REGION Network 46: Aviso 55 - El Secador Sullair 1 alcanzó la máxima cantidad de horas sin mantenimiento 2
   RUNG wire#powerrail
      Contact( "LimiteMantMS054_2" )
      Coil( "DB_ALA_PRE".x165 )
   END_RUNG
   // the same network as SCL:
   "DB_ALA_PRE".x165 := "LimiteMantMS054_2";
END_REGION

REGION Network 47: Aviso 56 - El Secador Sullair 2 alcanzó la máxima cantidad de horas sin mantenimiento 1
   RUNG wire#powerrail
      Contact( "LimiteMantMS055_1" )
      Coil( "DB_ALA_PRE".x166 )
   END_RUNG
   // the same network as SCL:
   "DB_ALA_PRE".x166 := "LimiteMantMS055_1";
END_REGION

REGION Network 48: Aviso 57 - El Secador Sullair 2 alcanzó la máxima cantidad de horas sin mantenimiento 2
   RUNG wire#powerrail
      Contact( "LimiteMantMS055_2" )
      Coil( "DB_ALA_PRE".x167 )
   END_RUNG
   // the same network as SCL:
   "DB_ALA_PRE".x167 := "LimiteMantMS055_2";
END_REGION

REGION Network 49: Aviso 58 - El Compresor Sullair 2 alcanzó la máxima cantidad de horas sin mantenimiento 1
   RUNG wire#powerrail
      Contact( "LimiteMantMC060_1" )
      Coil( "DB_ALA_PRE".x168 )
   END_RUNG
   // the same network as SCL:
   "DB_ALA_PRE".x168 := "LimiteMantMC060_1";
END_REGION

REGION Network 50: Aviso 59 - El Compresor Sullair 2 alcanzó la máxima cantidad de horas sin mantenimiento 2
   RUNG wire#powerrail
      Contact( "LimiteMantMC060_2" )
      Coil( "DB_ALA_PRE".x169 )
   END_RUNG
   // the same network as SCL:
   "DB_ALA_PRE".x169 := "LimiteMantMC060_2";
END_REGION

REGION Network 51: Aviso 60 - El Compresor Sullair 2 alcanzó la máxima cantidad de horas sin mantenimiento 3
   RUNG wire#powerrail
      Contact( "LimiteMantMC060_3" )
      Coil( "DB_ALA_PRE".x170 )
   END_RUNG
   // the same network as SCL:
   "DB_ALA_PRE".x170 := "LimiteMantMC060_3";
END_REGION

REGION Network 52: Aviso 61 - El Compresor Sullair 2 alcanzó la máxima cantidad de horas sin mantenimiento 4
   RUNG wire#powerrail
      Contact( "LimiteMantMC060_4" )
      Coil( "DB_ALA_PRE".x171 )
   END_RUNG
   // the same network as SCL:
   "DB_ALA_PRE".x171 := "LimiteMantMC060_4";
END_REGION

REGION Network 53: Aviso 62 - El Compresor Sullair 2 alcanzó la máxima cantidad de horas sin mantenimiento 5
   RUNG wire#powerrail
      Contact( "LimiteMantMC060_5" )
      Coil( "DB_ALA_PRE".x172 )
   END_RUNG
   // the same network as SCL:
   "DB_ALA_PRE".x172 := "LimiteMantMC060_5";
END_REGION

REGION Network 54: Aviso 63 - El Compresor Sullair 1 alcanzó la máxima cantidad de horas sin mantenimiento 1
   RUNG wire#powerrail
      Contact( "LimiteMantMC061_1" )
      Coil( "DB_ALA_PRE".x173 )
   END_RUNG
   // the same network as SCL:
   "DB_ALA_PRE".x173 := "LimiteMantMC061_1";
END_REGION

REGION Network 55: Aviso 64 - El Compresor Sullair 1 alcanzó la máxima cantidad de horas sin mantenimiento 2
   RUNG wire#powerrail
      Contact( "LimiteMantMC061_2" )
      Coil( "DB_ALA_PRE".x174 )
   END_RUNG
   // the same network as SCL:
   "DB_ALA_PRE".x174 := "LimiteMantMC061_2";
END_REGION

REGION Network 56: Aviso 65 - El Compresor Sullair 1 alcanzó la máxima cantidad de horas sin mantenimiento 3
   RUNG wire#powerrail
      Contact( "LimiteMantMC061_3" )
      Coil( "DB_ALA_PRE".x175 )
   END_RUNG
   // the same network as SCL:
   "DB_ALA_PRE".x175 := "LimiteMantMC061_3";
END_REGION

REGION Network 57: Aviso 84 - El Compresor Sullair 1 alcanzó la máxima cantidad de horas sin mantenimiento 4
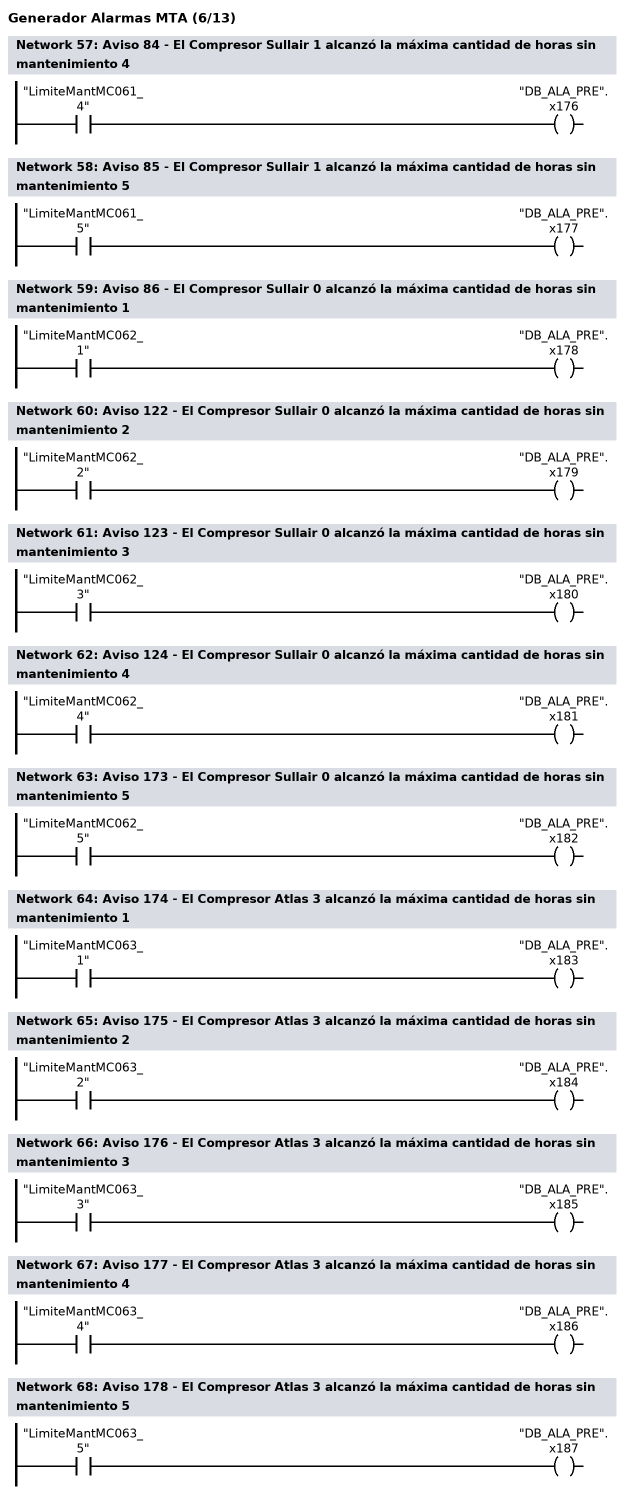
   RUNG wire#powerrail
      Contact( "LimiteMantMC061_4" )
      Coil( "DB_ALA_PRE".x176 )
   END_RUNG
   // the same network as SCL:
   "DB_ALA_PRE".x176 := "LimiteMantMC061_4";
END_REGION

REGION Network 58: Aviso 85 - El Compresor Sullair 1 alcanzó la máxima cantidad de horas sin mantenimiento 5
   RUNG wire#powerrail
      Contact( "LimiteMantMC061_5" )
      Coil( "DB_ALA_PRE".x177 )
   END_RUNG
   // the same network as SCL:
   "DB_ALA_PRE".x177 := "LimiteMantMC061_5";
END_REGION

REGION Network 59: Aviso 86 - El Compresor Sullair 0 alcanzó la máxima cantidad de horas sin mantenimiento 1
   RUNG wire#powerrail
      Contact( "LimiteMantMC062_1" )
      Coil( "DB_ALA_PRE".x178 )
   END_RUNG
   // the same network as SCL:
   "DB_ALA_PRE".x178 := "LimiteMantMC062_1";
END_REGION

REGION Network 60: Aviso 122 - El Compresor Sullair 0 alcanzó la máxima cantidad de horas sin mantenimiento 2
   RUNG wire#powerrail
      Contact( "LimiteMantMC062_2" )
      Coil( "DB_ALA_PRE".x179 )
   END_RUNG
   // the same network as SCL:
   "DB_ALA_PRE".x179 := "LimiteMantMC062_2";
END_REGION

REGION Network 61: Aviso 123 - El Compresor Sullair 0 alcanzó la máxima cantidad de horas sin mantenimiento 3
   RUNG wire#powerrail
      Contact( "LimiteMantMC062_3" )
      Coil( "DB_ALA_PRE".x180 )
   END_RUNG
   // the same network as SCL:
   "DB_ALA_PRE".x180 := "LimiteMantMC062_3";
END_REGION

REGION Network 62: Aviso 124 - El Compresor Sullair 0 alcanzó la máxima cantidad de horas sin mantenimiento 4
   RUNG wire#powerrail
      Contact( "LimiteMantMC062_4" )
      Coil( "DB_ALA_PRE".x181 )
   END_RUNG
   // the same network as SCL:
   "DB_ALA_PRE".x181 := "LimiteMantMC062_4";
END_REGION

REGION Network 63: Aviso 173 - El Compresor Sullair 0 alcanzó la máxima cantidad de horas sin mantenimiento 5
   RUNG wire#powerrail
      Contact( "LimiteMantMC062_5" )
      Coil( "DB_ALA_PRE".x182 )
   END_RUNG
   // the same network as SCL:
   "DB_ALA_PRE".x182 := "LimiteMantMC062_5";
END_REGION

REGION Network 64: Aviso 174 - El Compresor Atlas 3 alcanzó la máxima cantidad de horas sin mantenimiento 1
   RUNG wire#powerrail
      Contact( "LimiteMantMC063_1" )
      Coil( "DB_ALA_PRE".x183 )
   END_RUNG
   // the same network as SCL:
   "DB_ALA_PRE".x183 := "LimiteMantMC063_1";
END_REGION

REGION Network 65: Aviso 175 - El Compresor Atlas 3 alcanzó la máxima cantidad de horas sin mantenimiento 2
   RUNG wire#powerrail
      Contact( "LimiteMantMC063_2" )
      Coil( "DB_ALA_PRE".x184 )
   END_RUNG
   // the same network as SCL:
   "DB_ALA_PRE".x184 := "LimiteMantMC063_2";
END_REGION

REGION Network 66: Aviso 176 - El Compresor Atlas 3 alcanzó la máxima cantidad de horas sin mantenimiento 3
   RUNG wire#powerrail
      Contact( "LimiteMantMC063_3" )
      Coil( "DB_ALA_PRE".x185 )
   END_RUNG
   // the same network as SCL:
   "DB_ALA_PRE".x185 := "LimiteMantMC063_3";
END_REGION

REGION Network 67: Aviso 177 - El Compresor Atlas 3 alcanzó la máxima cantidad de horas sin mantenimiento 4
   RUNG wire#powerrail
      Contact( "LimiteMantMC063_4" )
      Coil( "DB_ALA_PRE".x186 )
   END_RUNG
   // the same network as SCL:
   "DB_ALA_PRE".x186 := "LimiteMantMC063_4";
END_REGION

REGION Network 68: Aviso 178 - El Compresor Atlas 3 alcanzó la máxima cantidad de horas sin mantenimiento 5
   RUNG wire#powerrail
      Contact( "LimiteMantMC063_5" )
      Coil( "DB_ALA_PRE".x187 )
   END_RUNG
   // the same network as SCL:
   "DB_ALA_PRE".x187 := "LimiteMantMC063_5";
END_REGION

REGION Network 69: Aviso 179 - El Compresor Atlas 2 alcanzó la máxima cantidad de horas sin mantenimiento 1
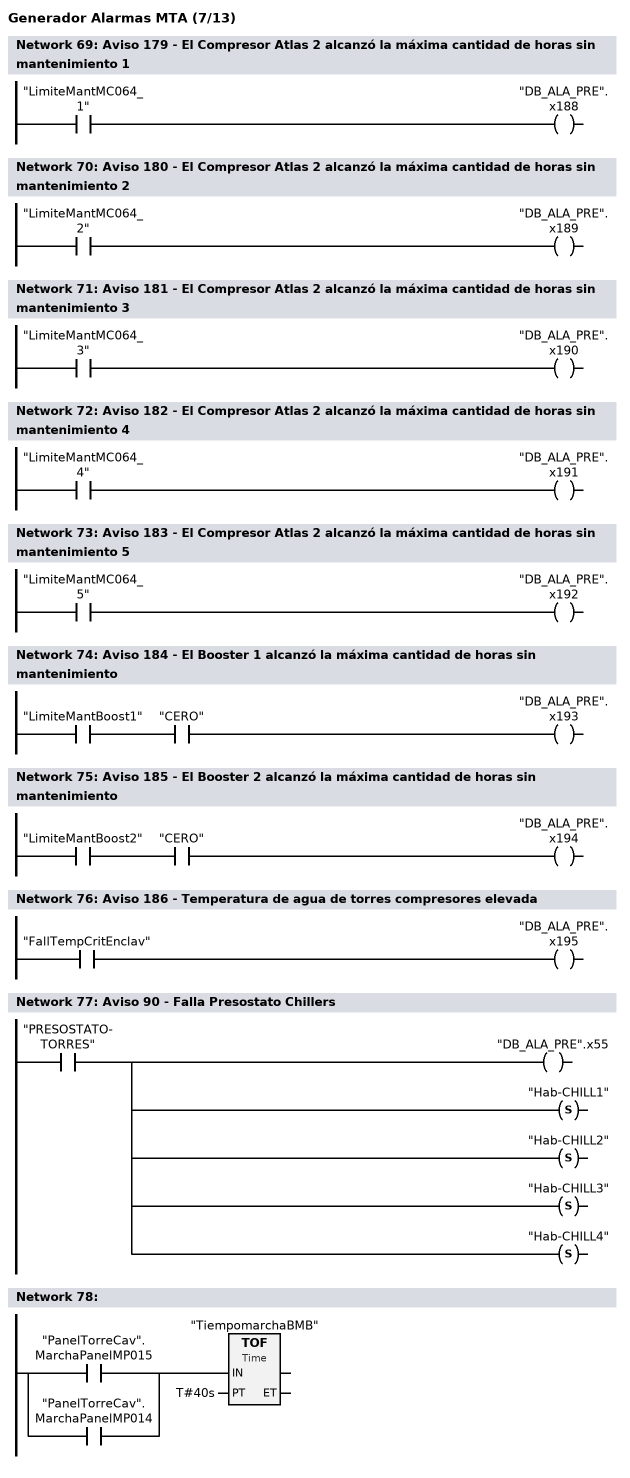
   RUNG wire#powerrail
      Contact( "LimiteMantMC064_1" )
      Coil( "DB_ALA_PRE".x188 )
   END_RUNG
   // the same network as SCL:
   "DB_ALA_PRE".x188 := "LimiteMantMC064_1";
END_REGION

REGION Network 70: Aviso 180 - El Compresor Atlas 2 alcanzó la máxima cantidad de horas sin mantenimiento 2
   RUNG wire#powerrail
      Contact( "LimiteMantMC064_2" )
      Coil( "DB_ALA_PRE".x189 )
   END_RUNG
   // the same network as SCL:
   "DB_ALA_PRE".x189 := "LimiteMantMC064_2";
END_REGION

REGION Network 71: Aviso 181 - El Compresor Atlas 2 alcanzó la máxima cantidad de horas sin mantenimiento 3
   RUNG wire#powerrail
      Contact( "LimiteMantMC064_3" )
      Coil( "DB_ALA_PRE".x190 )
   END_RUNG
   // the same network as SCL:
   "DB_ALA_PRE".x190 := "LimiteMantMC064_3";
END_REGION

REGION Network 72: Aviso 182 - El Compresor Atlas 2 alcanzó la máxima cantidad de horas sin mantenimiento 4
   RUNG wire#powerrail
      Contact( "LimiteMantMC064_4" )
      Coil( "DB_ALA_PRE".x191 )
   END_RUNG
   // the same network as SCL:
   "DB_ALA_PRE".x191 := "LimiteMantMC064_4";
END_REGION

REGION Network 73: Aviso 183 - El Compresor Atlas 2 alcanzó la máxima cantidad de horas sin mantenimiento 5
   RUNG wire#powerrail
      Contact( "LimiteMantMC064_5" )
      Coil( "DB_ALA_PRE".x192 )
   END_RUNG
   // the same network as SCL:
   "DB_ALA_PRE".x192 := "LimiteMantMC064_5";
END_REGION

REGION Network 74: Aviso 184 - El Booster 1 alcanzó la máxima cantidad de horas sin mantenimiento
   RUNG wire#powerrail
      Contact( "LimiteMantBoost1" )
      Contact( "CERO" )
      Coil( "DB_ALA_PRE".x193 )
   END_RUNG
   // the same network as SCL:
   "DB_ALA_PRE".x193 := "LimiteMantBoost1" AND "CERO";
END_REGION

REGION Network 75: Aviso 185 - El Booster 2 alcanzó la máxima cantidad de horas sin mantenimiento
   RUNG wire#powerrail
      Contact( "LimiteMantBoost2" )
      Contact( "CERO" )
      Coil( "DB_ALA_PRE".x194 )
   END_RUNG
   // the same network as SCL:
   "DB_ALA_PRE".x194 := "LimiteMantBoost2" AND "CERO";
END_REGION

REGION Network 76: Aviso 186 - Temperatura de agua de torres compresores elevada
   RUNG wire#powerrail
      Contact( "FallTempCritEnclav" )
      Coil( "DB_ALA_PRE".x195 )
   END_RUNG
   // the same network as SCL:
   "DB_ALA_PRE".x195 := "FallTempCritEnclav";
END_REGION

REGION Network 77: Aviso 90 - Falla Presostato Chillers
   RUNG wire#powerrail
      Contact( "PRESOSTATO-TORRES" )
      wire#w1
      Coil( "DB_ALA_PRE".x55 )
   END_RUNG
   RUNG wire#w1
      S_Coil( "Hab-CHILL1" )
   END_RUNG
   RUNG wire#w1
      S_Coil( "Hab-CHILL2" )
   END_RUNG
   RUNG wire#w1
      S_Coil( "Hab-CHILL3" )
   END_RUNG
   RUNG wire#w1
      S_Coil( "Hab-CHILL4" )
   END_RUNG
   // the same network as SCL:
   "DB_ALA_PRE".x55 := "PRESOSTATO-TORRES";
   IF "PRESOSTATO-TORRES" THEN
       "Hab-CHILL1" := TRUE;
       "Hab-CHILL2" := TRUE;
       "Hab-CHILL3" := TRUE;
       "Hab-CHILL4" := TRUE;
   END_IF;
END_REGION

REGION Network 78
   "TiempomarchaBMB".TOF(IN := "PanelTorreCav".MarchaPanelMP015 OR "PanelTorreCav".MarchaPanelMP014,
                         PT := T#40s);
END_REGION

REGION Network 79
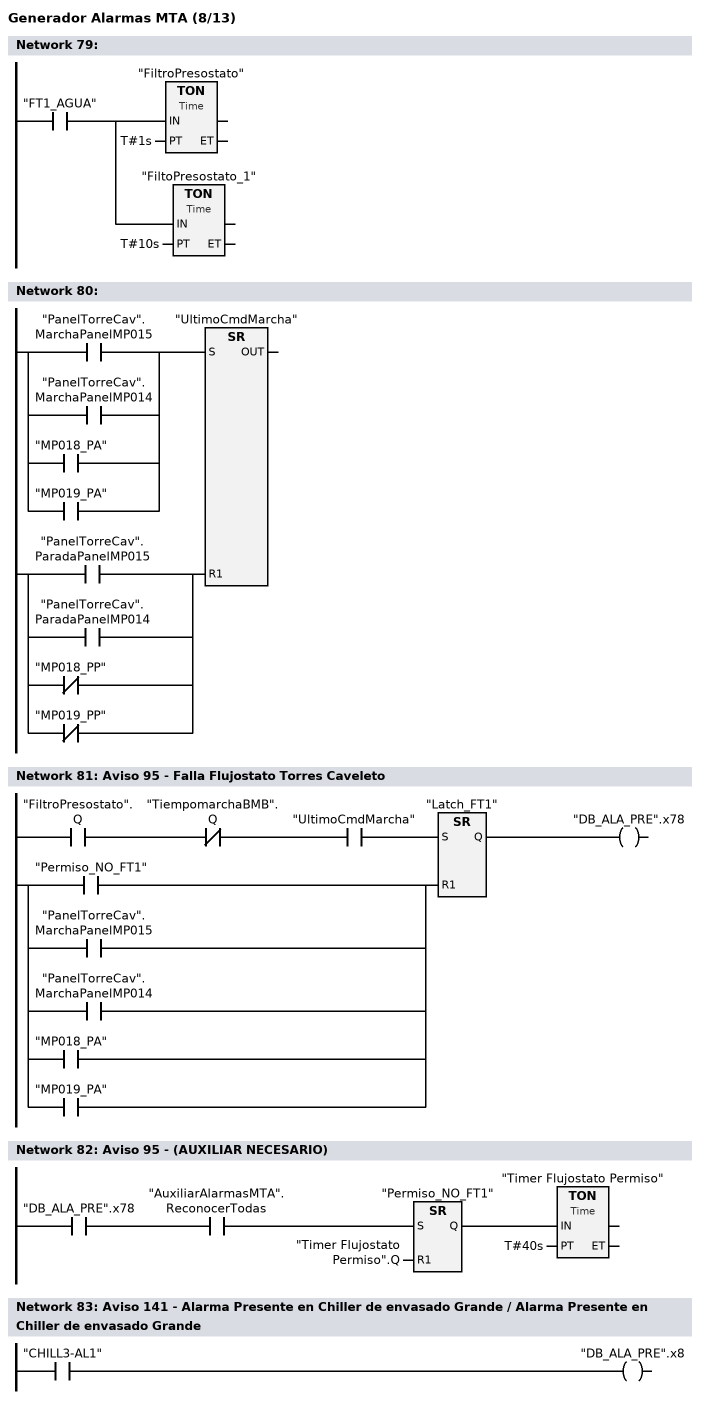
   "FiltroPresostato".TON(IN := "FT1_AGUA", PT := T#1s);
   "FiltoPresostato_1".TON(IN := "FT1_AGUA", PT := T#10s);
END_REGION

REGION Network 80
   RUNG wire#powerrail
      Contact( "PanelTorreCav".MarchaPanelMP015 )
      wire#w1
      S_SR(operand := "UltimoCmdMarcha", r1 := wire#w2)
   END_RUNG
   RUNG wire#powerrail
      Contact( "PanelTorreCav".MarchaPanelMP014 )
   END_RUNG wire#w1
   RUNG wire#powerrail
      Contact( "MP018_PA" )
   END_RUNG wire#w1
   RUNG wire#powerrail
      Contact( "MP019_PA" )
   END_RUNG wire#w1
   RUNG wire#powerrail
      Contact( "PanelTorreCav".ParadaPanelMP015 )
   END_RUNG wire#w2
   RUNG wire#powerrail
      Contact( "PanelTorreCav".ParadaPanelMP014 )
   END_RUNG wire#w2
   RUNG wire#powerrail
      I_Contact( "MP018_PP" )
   END_RUNG wire#w2
   RUNG wire#powerrail
      I_Contact( "MP019_PP" )
   END_RUNG wire#w2
   // the same network as SCL:
   IF "PanelTorreCav".MarchaPanelMP015 OR "PanelTorreCav".MarchaPanelMP014 OR "MP018_PA" OR "MP019_PA" THEN
       "UltimoCmdMarcha" := TRUE;   // SR flip-flop
   END_IF;
   IF "PanelTorreCav".ParadaPanelMP015 OR "PanelTorreCav".ParadaPanelMP014 OR NOT "MP018_PP" OR NOT "MP019_PP" THEN
       "UltimoCmdMarcha" := FALSE;
   END_IF;
END_REGION

REGION Network 81: Aviso 95 - Falla Flujostato Torres Caveleto
   RUNG wire#powerrail
      Contact( "FiltroPresostato".Q )
      I_Contact( "TiempomarchaBMB".Q )
      Contact( "UltimoCmdMarcha" )
      S_SR(operand := "Latch_FT1", r1 := wire#w1)
      Coil( "DB_ALA_PRE".x78 )
   END_RUNG
   RUNG wire#powerrail
      Contact( "Permiso_NO_FT1" )
   END_RUNG wire#w1
   RUNG wire#powerrail
      Contact( "PanelTorreCav".MarchaPanelMP015 )
   END_RUNG wire#w1
   RUNG wire#powerrail
      Contact( "PanelTorreCav".MarchaPanelMP014 )
   END_RUNG wire#w1
   RUNG wire#powerrail
      Contact( "MP018_PA" )
   END_RUNG wire#w1
   RUNG wire#powerrail
      Contact( "MP019_PA" )
   END_RUNG wire#w1
   // the same network as SCL:
   IF "FiltroPresostato".Q AND NOT "TiempomarchaBMB".Q AND "UltimoCmdMarcha" THEN
       "Latch_FT1" := TRUE;   // SR flip-flop
   END_IF;
   IF "Permiso_NO_FT1" OR "PanelTorreCav".MarchaPanelMP015 OR "PanelTorreCav".MarchaPanelMP014 OR "MP018_PA" OR "MP019_PA" THEN
       "Latch_FT1" := FALSE;
   END_IF;
   "DB_ALA_PRE".x78 := "Latch_FT1";
END_REGION

REGION Network 82: Aviso 95 - (AUXILIAR NECESARIO)
   IF "DB_ALA_PRE".x78 AND "AuxiliarAlarmasMTA".ReconocerTodas THEN
       "Permiso_NO_FT1" := TRUE;   // SR flip-flop
   END_IF;
   IF "Timer Flujostato Permiso".Q THEN "Permiso_NO_FT1" := FALSE; END_IF;
   "Timer Flujostato Permiso".TON(IN := "Permiso_NO_FT1", PT := T#40s);
END_REGION

REGION Network 83: Aviso 141 - Alarma Presente en Chiller de envasado Grande / Alarma Presente en Chiller de envasado Grande
   RUNG wire#powerrail
      Contact( "CHILL3-AL1" )
      Coil( "DB_ALA_PRE".x8 )
   END_RUNG
   // the same network as SCL:
   "DB_ALA_PRE".x8 := "CHILL3-AL1";
END_REGION

REGION Network 84: Aviso 142 - Alarma Presente en Chiller de soplado Grande
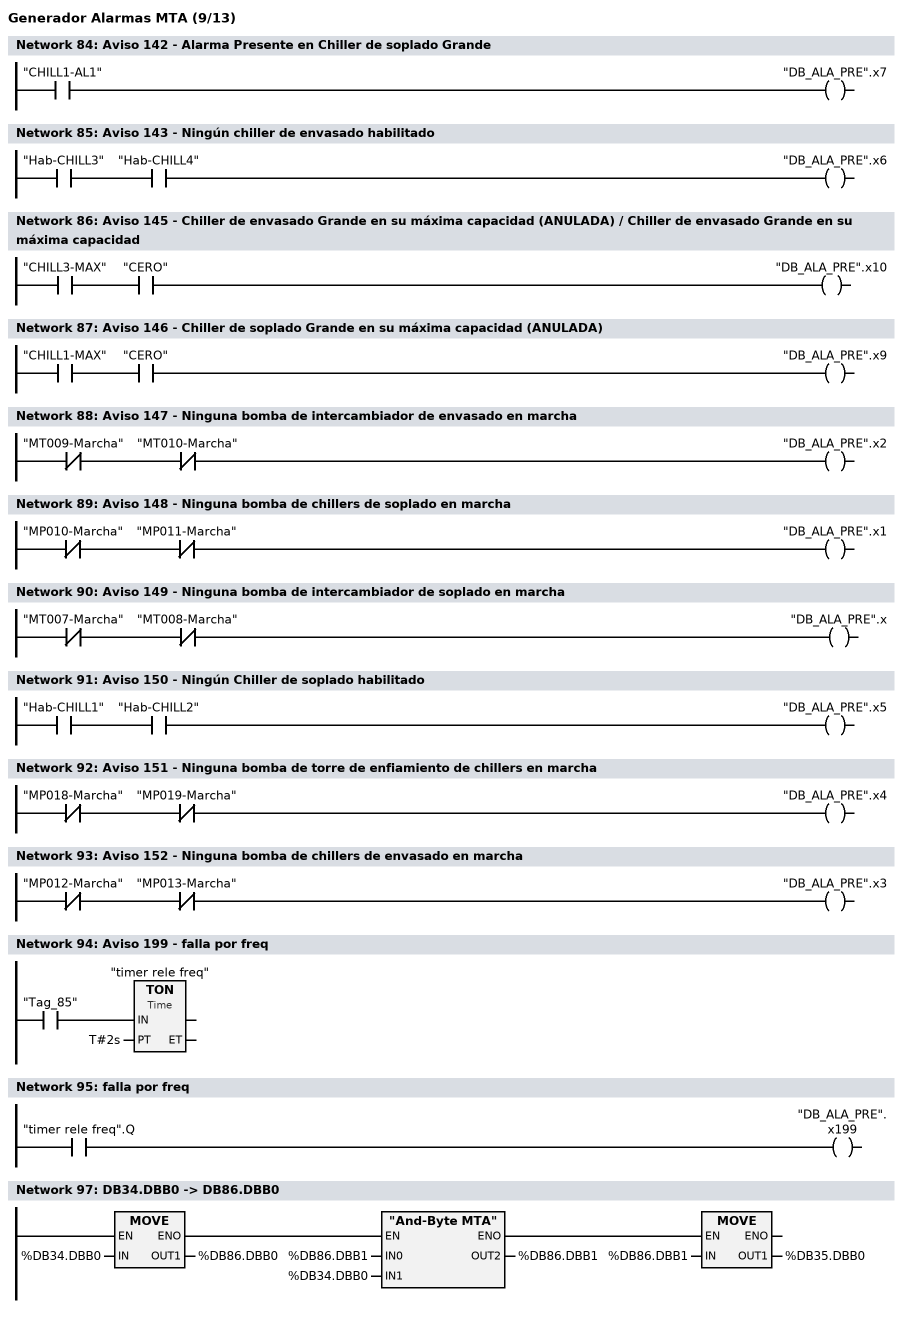
   RUNG wire#powerrail
      Contact( "CHILL1-AL1" )
      Coil( "DB_ALA_PRE".x7 )
   END_RUNG
   // the same network as SCL:
   "DB_ALA_PRE".x7 := "CHILL1-AL1";
END_REGION

REGION Network 85: Aviso 143 - Ningún chiller de envasado habilitado
   RUNG wire#powerrail
      Contact( "Hab-CHILL3" )
      Contact( "Hab-CHILL4" )
      Coil( "DB_ALA_PRE".x6 )
   END_RUNG
   // the same network as SCL:
   "DB_ALA_PRE".x6 := "Hab-CHILL3" AND "Hab-CHILL4";
END_REGION

REGION Network 86: Aviso 145 - Chiller de envasado Grande en su máxima capacidad (ANULADA) / Chiller de envasado Grande en su máxima capacidad
   RUNG wire#powerrail
      Contact( "CHILL3-MAX" )
      Contact( "CERO" )
      Coil( "DB_ALA_PRE".x10 )
   END_RUNG
   // the same network as SCL:
   "DB_ALA_PRE".x10 := "CHILL3-MAX" AND "CERO";
END_REGION

REGION Network 87: Aviso 146 - Chiller de soplado Grande en su máxima capacidad (ANULADA)
   RUNG wire#powerrail
      Contact( "CHILL1-MAX" )
      Contact( "CERO" )
      Coil( "DB_ALA_PRE".x9 )
   END_RUNG
   // the same network as SCL:
   "DB_ALA_PRE".x9 := "CHILL1-MAX" AND "CERO";
END_REGION

REGION Network 88: Aviso 147 - Ninguna bomba de intercambiador de envasado en marcha
   RUNG wire#powerrail
      I_Contact( "MT009-Marcha" )
      I_Contact( "MT010-Marcha" )
      Coil( "DB_ALA_PRE".x2 )
   END_RUNG
   // the same network as SCL:
   "DB_ALA_PRE".x2 := NOT "MT009-Marcha" AND NOT "MT010-Marcha";
END_REGION

REGION Network 89: Aviso 148 - Ninguna bomba de chillers de soplado en marcha
   RUNG wire#powerrail
      I_Contact( "MP010-Marcha" )
      I_Contact( "MP011-Marcha" )
      Coil( "DB_ALA_PRE".x1 )
   END_RUNG
   // the same network as SCL:
   "DB_ALA_PRE".x1 := NOT "MP010-Marcha" AND NOT "MP011-Marcha";
END_REGION

REGION Network 90: Aviso 149 - Ninguna bomba de intercambiador de soplado en marcha
   RUNG wire#powerrail
      I_Contact( "MT007-Marcha" )
      I_Contact( "MT008-Marcha" )
      Coil( "DB_ALA_PRE".x )
   END_RUNG
   // the same network as SCL:
   "DB_ALA_PRE".x := NOT "MT007-Marcha" AND NOT "MT008-Marcha";
END_REGION

REGION Network 91: Aviso 150 - Ningún Chiller de soplado habilitado
   RUNG wire#powerrail
      Contact( "Hab-CHILL1" )
      Contact( "Hab-CHILL2" )
      Coil( "DB_ALA_PRE".x5 )
   END_RUNG
   // the same network as SCL:
   "DB_ALA_PRE".x5 := "Hab-CHILL1" AND "Hab-CHILL2";
END_REGION

REGION Network 92: Aviso 151 - Ninguna bomba de torre de enfiamiento de chillers en marcha
   RUNG wire#powerrail
      I_Contact( "MP018-Marcha" )
      I_Contact( "MP019-Marcha" )
      Coil( "DB_ALA_PRE".x4 )
   END_RUNG
   // the same network as SCL:
   "DB_ALA_PRE".x4 := NOT "MP018-Marcha" AND NOT "MP019-Marcha";
END_REGION

REGION Network 93: Aviso 152 - Ninguna bomba de chillers de envasado en marcha
   RUNG wire#powerrail
      I_Contact( "MP012-Marcha" )
      I_Contact( "MP013-Marcha" )
      Coil( "DB_ALA_PRE".x3 )
   END_RUNG
   // the same network as SCL:
   "DB_ALA_PRE".x3 := NOT "MP012-Marcha" AND NOT "MP013-Marcha";
END_REGION

REGION Network 94: Aviso 199 - falla por freq
   "timer rele freq".TON(IN := "Tag_85", PT := T#2s);
END_REGION

REGION Network 95: falla por freq
   RUNG wire#powerrail
      Contact( "timer rele freq".Q )
      Coil( "DB_ALA_PRE".x199 )
   END_RUNG
   // the same network as SCL:
   "DB_ALA_PRE".x199 := "timer rele freq".Q;
END_REGION

REGION Network 97: DB34.DBB0 -> DB86.DBB0
   RUNG wire#powerrail
      { S7_GenerateENO := "TRUE" } Move(in := %DB34.DBB0, out1 => %DB86.DBB0)
      "And-Byte MTA"(IN0 := %DB86.DBB1, IN1 := %DB34.DBB0, OUT2 => %DB86.DBB1)
      { S7_GenerateENO := "TRUE" } Move(in := %DB86.DBB1, out1 => %DB35.DBB0)
   END_RUNG
   // the same network as SCL:
   // ENO of a box is taken as its EN; it also drops when the box reports an error
   %DB86.DBB0 := %DB34.DBB0;
   "And-Byte MTA"(IN0 := %DB86.DBB1, IN1 := %DB34.DBB0, OUT2 => %DB86.DBB1, ENO => #_w1);
   IF #_w1 THEN %DB35.DBB0 := %DB86.DBB1; END_IF;
END_REGION

REGION Network 98: DB34.DBB1 -> DB86.DBB2 / 8 y 8
   // Alarma Presente en Chiller de envasado Grande
   // Chiller de soplado Grande en su máxima capacidad
   // Chiller de envasado Grande en su máxima capacidad
   // Falla Térmico MT007
   // Falla Contactor MT007
   // Falla Térmico MT008
   // Falla Contactor MT008
   // Falla Térmico MT009
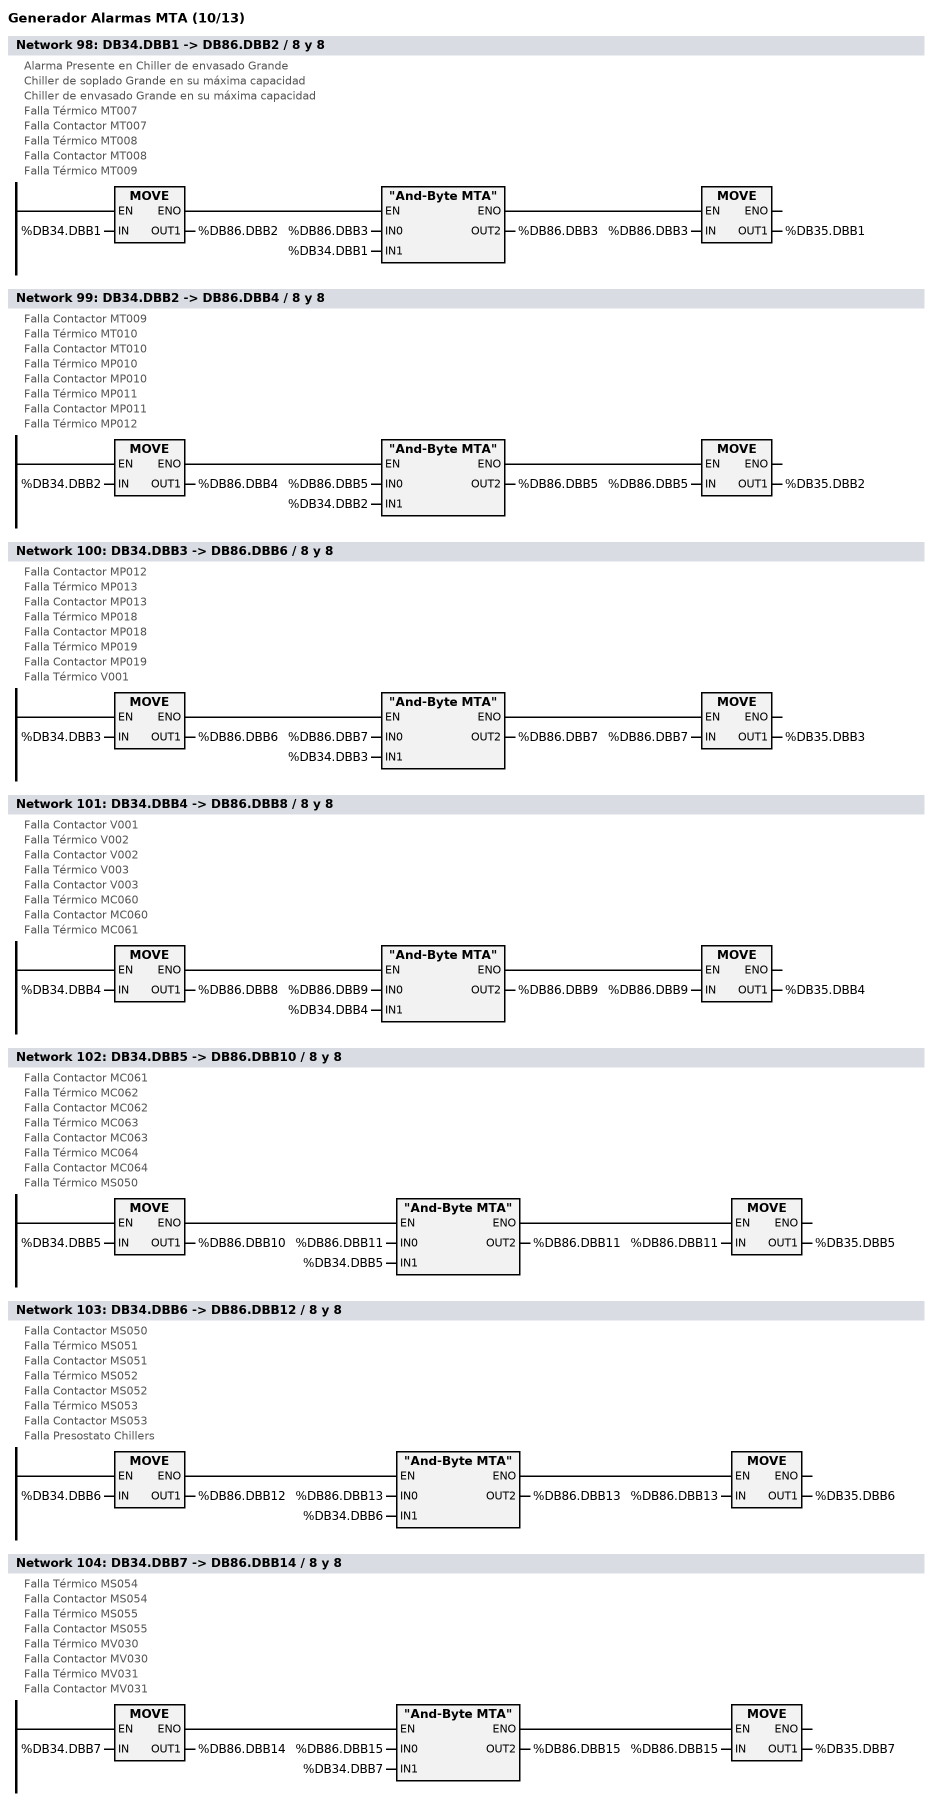
   RUNG wire#powerrail
      { S7_GenerateENO := "TRUE" } Move(in := %DB34.DBB1, out1 => %DB86.DBB2)
      "And-Byte MTA"(IN0 := %DB86.DBB3, IN1 := %DB34.DBB1, OUT2 => %DB86.DBB3)
      { S7_GenerateENO := "TRUE" } Move(in := %DB86.DBB3, out1 => %DB35.DBB1)
   END_RUNG
   // the same network as SCL:
   // ENO of a box is taken as its EN; it also drops when the box reports an error
   %DB86.DBB2 := %DB34.DBB1;
   "And-Byte MTA"(IN0 := %DB86.DBB3, IN1 := %DB34.DBB1, OUT2 => %DB86.DBB3, ENO => #_w1);
   IF #_w1 THEN %DB35.DBB1 := %DB86.DBB3; END_IF;
END_REGION

REGION Network 99: DB34.DBB2 -> DB86.DBB4 / 8 y 8
   // Falla Contactor MT009
   // Falla Térmico MT010
   // Falla Contactor MT010
   // Falla Térmico MP010
   // Falla Contactor MP010
   // Falla Térmico MP011
   // Falla Contactor MP011
   // Falla Térmico MP012
   RUNG wire#powerrail
      { S7_GenerateENO := "TRUE" } Move(in := %DB34.DBB2, out1 => %DB86.DBB4)
      "And-Byte MTA"(IN0 := %DB86.DBB5, IN1 := %DB34.DBB2, OUT2 => %DB86.DBB5)
      { S7_GenerateENO := "TRUE" } Move(in := %DB86.DBB5, out1 => %DB35.DBB2)
   END_RUNG
   // the same network as SCL:
   // ENO of a box is taken as its EN; it also drops when the box reports an error
   %DB86.DBB4 := %DB34.DBB2;
   "And-Byte MTA"(IN0 := %DB86.DBB5, IN1 := %DB34.DBB2, OUT2 => %DB86.DBB5, ENO => #_w1);
   IF #_w1 THEN %DB35.DBB2 := %DB86.DBB5; END_IF;
END_REGION

REGION Network 100: DB34.DBB3 -> DB86.DBB6 / 8 y 8
   // Falla Contactor MP012
   // Falla Térmico MP013
   // Falla Contactor MP013
   // Falla Térmico MP018
   // Falla Contactor MP018
   // Falla Térmico MP019
   // Falla Contactor MP019
   // Falla Térmico V001
   RUNG wire#powerrail
      { S7_GenerateENO := "TRUE" } Move(in := %DB34.DBB3, out1 => %DB86.DBB6)
      "And-Byte MTA"(IN0 := %DB86.DBB7, IN1 := %DB34.DBB3, OUT2 => %DB86.DBB7)
      { S7_GenerateENO := "TRUE" } Move(in := %DB86.DBB7, out1 => %DB35.DBB3)
   END_RUNG
   // the same network as SCL:
   // ENO of a box is taken as its EN; it also drops when the box reports an error
   %DB86.DBB6 := %DB34.DBB3;
   "And-Byte MTA"(IN0 := %DB86.DBB7, IN1 := %DB34.DBB3, OUT2 => %DB86.DBB7, ENO => #_w1);
   IF #_w1 THEN %DB35.DBB3 := %DB86.DBB7; END_IF;
END_REGION

REGION Network 101: DB34.DBB4 -> DB86.DBB8 / 8 y 8
   // Falla Contactor V001
   // Falla Térmico V002
   // Falla Contactor V002
   // Falla Térmico V003
   // Falla Contactor V003
   // Falla Térmico MC060
   // Falla Contactor MC060
   // Falla Térmico MC061
   RUNG wire#powerrail
      { S7_GenerateENO := "TRUE" } Move(in := %DB34.DBB4, out1 => %DB86.DBB8)
      "And-Byte MTA"(IN0 := %DB86.DBB9, IN1 := %DB34.DBB4, OUT2 => %DB86.DBB9)
      { S7_GenerateENO := "TRUE" } Move(in := %DB86.DBB9, out1 => %DB35.DBB4)
   END_RUNG
   // the same network as SCL:
   // ENO of a box is taken as its EN; it also drops when the box reports an error
   %DB86.DBB8 := %DB34.DBB4;
   "And-Byte MTA"(IN0 := %DB86.DBB9, IN1 := %DB34.DBB4, OUT2 => %DB86.DBB9, ENO => #_w1);
   IF #_w1 THEN %DB35.DBB4 := %DB86.DBB9; END_IF;
END_REGION

REGION Network 102: DB34.DBB5 -> DB86.DBB10 / 8 y 8
   // Falla Contactor MC061
   // Falla Térmico MC062
   // Falla Contactor MC062
   // Falla Térmico MC063
   // Falla Contactor MC063
   // Falla Térmico MC064
   // Falla Contactor MC064
   // Falla Térmico MS050
   RUNG wire#powerrail
      { S7_GenerateENO := "TRUE" } Move(in := %DB34.DBB5, out1 => %DB86.DBB10)
      "And-Byte MTA"(IN0 := %DB86.DBB11, IN1 := %DB34.DBB5, OUT2 => %DB86.DBB11)
      { S7_GenerateENO := "TRUE" } Move(in := %DB86.DBB11, out1 => %DB35.DBB5)
   END_RUNG
   // the same network as SCL:
   // ENO of a box is taken as its EN; it also drops when the box reports an error
   %DB86.DBB10 := %DB34.DBB5;
   "And-Byte MTA"(IN0 := %DB86.DBB11, IN1 := %DB34.DBB5, OUT2 => %DB86.DBB11, ENO => #_w1);
   IF #_w1 THEN %DB35.DBB5 := %DB86.DBB11; END_IF;
END_REGION

REGION Network 103: DB34.DBB6 -> DB86.DBB12 / 8 y 8
   // Falla Contactor MS050
   // Falla Térmico MS051
   // Falla Contactor MS051
   // Falla Térmico MS052
   // Falla Contactor MS052
   // Falla Térmico MS053
   // Falla Contactor MS053
   // Falla Presostato Chillers
   RUNG wire#powerrail
      { S7_GenerateENO := "TRUE" } Move(in := %DB34.DBB6, out1 => %DB86.DBB12)
      "And-Byte MTA"(IN0 := %DB86.DBB13, IN1 := %DB34.DBB6, OUT2 => %DB86.DBB13)
      { S7_GenerateENO := "TRUE" } Move(in := %DB86.DBB13, out1 => %DB35.DBB6)
   END_RUNG
   // the same network as SCL:
   // ENO of a box is taken as its EN; it also drops when the box reports an error
   %DB86.DBB12 := %DB34.DBB6;
   "And-Byte MTA"(IN0 := %DB86.DBB13, IN1 := %DB34.DBB6, OUT2 => %DB86.DBB13, ENO => #_w1);
   IF #_w1 THEN %DB35.DBB6 := %DB86.DBB13; END_IF;
END_REGION

REGION Network 104: DB34.DBB7 -> DB86.DBB14 / 8 y 8
   // Falla Térmico MS054
   // Falla Contactor MS054
   // Falla Térmico MS055
   // Falla Contactor MS055
   // Falla Térmico MV030
   // Falla Contactor MV030
   // Falla Térmico MV031
   // Falla Contactor MV031
   RUNG wire#powerrail
      { S7_GenerateENO := "TRUE" } Move(in := %DB34.DBB7, out1 => %DB86.DBB14)
      "And-Byte MTA"(IN0 := %DB86.DBB15, IN1 := %DB34.DBB7, OUT2 => %DB86.DBB15)
      { S7_GenerateENO := "TRUE" } Move(in := %DB86.DBB15, out1 => %DB35.DBB7)
   END_RUNG
   // the same network as SCL:
   // ENO of a box is taken as its EN; it also drops when the box reports an error
   %DB86.DBB14 := %DB34.DBB7;
   "And-Byte MTA"(IN0 := %DB86.DBB15, IN1 := %DB34.DBB7, OUT2 => %DB86.DBB15, ENO => #_w1);
   IF #_w1 THEN %DB35.DBB7 := %DB86.DBB15; END_IF;
END_REGION

REGION Network 105: DB34.DBB8 -> DB86.DBB16 / 8 y 8
   // Falla Térmico MP014
   // Falla Contactor MP014
   // Falla Térmico MP015
   // Falla Contactor MP015
   // Falla Térmico MC001
   // Falla Contactor MC001
   // Falla Térmico MC002
   // Falla Contactor MC002
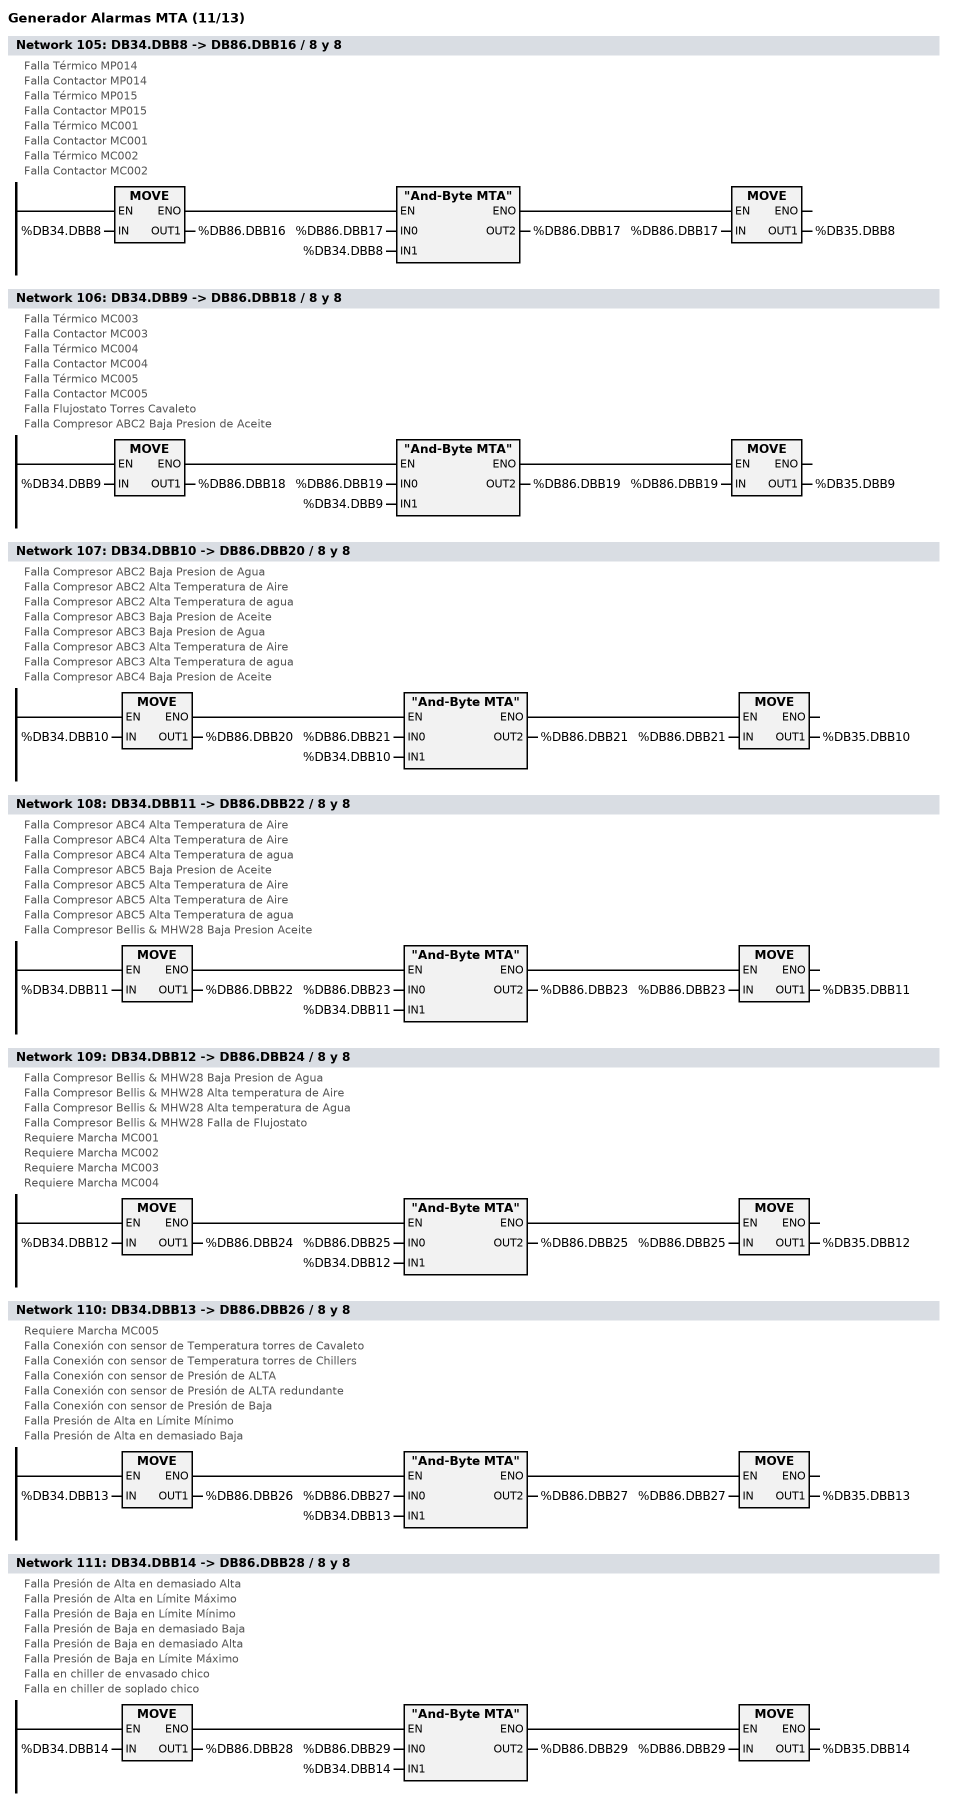
   RUNG wire#powerrail
      { S7_GenerateENO := "TRUE" } Move(in := %DB34.DBB8, out1 => %DB86.DBB16)
      "And-Byte MTA"(IN0 := %DB86.DBB17, IN1 := %DB34.DBB8, OUT2 => %DB86.DBB17)
      { S7_GenerateENO := "TRUE" } Move(in := %DB86.DBB17, out1 => %DB35.DBB8)
   END_RUNG
   // the same network as SCL:
   // ENO of a box is taken as its EN; it also drops when the box reports an error
   %DB86.DBB16 := %DB34.DBB8;
   "And-Byte MTA"(IN0 := %DB86.DBB17, IN1 := %DB34.DBB8, OUT2 => %DB86.DBB17, ENO => #_w1);
   IF #_w1 THEN %DB35.DBB8 := %DB86.DBB17; END_IF;
END_REGION

REGION Network 106: DB34.DBB9 -> DB86.DBB18 / 8 y 8
   // Falla Térmico MC003
   // Falla Contactor MC003
   // Falla Térmico MC004
   // Falla Contactor MC004
   // Falla Térmico MC005
   // Falla Contactor MC005
   // Falla Flujostato Torres Cavaleto
   // Falla Compresor ABC2 Baja Presion de Aceite
   RUNG wire#powerrail
      { S7_GenerateENO := "TRUE" } Move(in := %DB34.DBB9, out1 => %DB86.DBB18)
      "And-Byte MTA"(IN0 := %DB86.DBB19, IN1 := %DB34.DBB9, OUT2 => %DB86.DBB19)
      { S7_GenerateENO := "TRUE" } Move(in := %DB86.DBB19, out1 => %DB35.DBB9)
   END_RUNG
   // the same network as SCL:
   // ENO of a box is taken as its EN; it also drops when the box reports an error
   %DB86.DBB18 := %DB34.DBB9;
   "And-Byte MTA"(IN0 := %DB86.DBB19, IN1 := %DB34.DBB9, OUT2 => %DB86.DBB19, ENO => #_w1);
   IF #_w1 THEN %DB35.DBB9 := %DB86.DBB19; END_IF;
END_REGION
